VERSION : 0.0
   STRUCT
      doMotorOn : Bool;   // Systemoutput: Status for Motor OFF
      doMotorOff : Bool;   // Systemoutput: Status for Motor ON
      doCycleOn : Bool;   // Systemoutput: Robotprogram is running
      doIRBinAuto : Bool;   // Systemoutput: Robot is in operationmode AUTO
      doSysError : Bool;   // Systemoutput: Robot has an systemerror
      doEmStop_Akt : Bool;   // Systemoutput: Emergencystop at robot is active
      doMot_On_OK : Bool;   // Systemoutput: Automaticstopcicuites are OK
      do01_008 : Bool;   // Spare
      doIRBInHome : Bool;   // Worldzoneoutput: Robot is in Homeposition
      doIRBInMaintP : Bool;   // Worldzoneoutput: Robot is in Maintenanceposition
      doIRBOutRange : Bool;   // Worldzoneoutput: Robot near the end of it´s workingarealimitation
      doIRBOutRangMC : Bool;   // Worldzoneoutput: Robot is out of the mould
      doIRBOutRanMC1 : Bool;   // Worldzoneoutput: Robot is outside the mould carrier 1
      doIRBOutRanMC2 : Bool;   // Worldzoneoutput: Robot is outside the mould carrier 2
      doIRBOutRanMC3 : Bool;   // Worldzoneoutput: Robot is outside the mould carrier 3
      doIRBOutRanMC4 : Bool;   // Worldzoneoutput: Robot is outside the mould carrier 4
      doCycleStarted : Bool;   // The programcycle is startet
      doCycleEnd : Bool;   // The programcycle is finished
      doProgNoReaded : Bool;   // The programnumber is readed
      doShotDigOut : Bool;   // 1st digital Shotware output // Signal to open the mixinghead
      doStopFormPLC : Bool;   // Signal to stop the foaming because the robotprogram has stoped
      doShotBreak : Bool;
      doCloseMould : Bool;   // Signal that the robot is out of the mould
      doCP_forward : Bool;
      doIRBInMaintP2 : Bool;   // Worldzoneoutput: Robot is in 2. Maintenanceposition
      do01_026 : Bool;   // Spare
      doIRBSyncWobj : Bool;   // The robot is synchronized (Tracking)
      doRobWaitWobj : Bool;   // The robot is waiting for synchronizes (Tracking)
      doInPosTeach : Bool;   // The robot is in the position to teaching
      doConveyorStopped : Bool;   // The conveyor is stop
      doZeroSpeed : Bool;   // Systemoutput: Conveyer is not moving
      do01_032 : Bool;   // Spare
      do01_033 : Bool;   // Spare
      doSafetyControlPos : Bool;   // Signal to control the synchronization position
      doSafetySynchronized : Bool;   // Signal from Robot EPS is synchronize
      doSafetySyncSwitch : Bool;   // Signal from Robot sync switch is actuated
      doSafetyArea_1 : Bool;   // 1 Safe Output Safe move / EPS
      doSafetyArea_2 : Bool;   // 2 Safe Output Safe move / EPS
      doSafetyArea_3 : Bool;   // 3 Safe Output Safe move / EPS
      doSafetyArea_4 : Bool;   // 4 Safe Output Safe move / EPS
      doSafetyArea_5 : Bool;   // 5 Safe Output Safe move / EPS
      doSafetyArea_6 : Bool;   // 6 Safe Output Safe move / EPS
      doSafetyArea_7 : Bool;   // 7 Safe Output Safe move / EPS
      doSafetyArea_8 : Bool;   // 8 Safe Output Safe move / EPS
      doSafetyPreWarn : Bool;   // Signal from pre warning robot sync
      doSafeZoneActiv : Bool;   // Robot is inside of a safe tool zone
      do01_047 : Bool;   // Spare
      doClose_Mould_1 : Bool;
      doClose_Mould_2 : Bool;
      doClose_Mould_3 : Bool;
      doClose_Mould_4 : Bool;
      doIRBinSprayP : Bool;
      doSprayValveOn : Bool;
      doStartSpray : Bool;
      doSprayEnd : Bool;
      doInWaitPos : Bool;   // Signal robot is waiting in teh waiting position
      doIRBInWaitP : Bool;   // Signal robot is waiting in teh waiting position // Cube
      do01_058 : Bool;   // Spare
      do01_059 : Bool;   // Spare
      doCleaningPLC : Bool;   // Control the mixinghead cleaner or a brush station
      doCleanOsziJet : Bool;   // Control the air for blow out the oszilation holes
      doBlowAir : Bool;   // Control the air for blow inside the mixinghead
      doCleanBrushOn : Bool;   // Control the cleaning for the mixinghead
      doFlushing : Bool;
      doInFlushposSpray : Bool;
      doShotDigOut2 : Bool;   // 2nd digital Shotware output
      doShotDigOut3 : Bool;   // 3rd digital Shotware output
      do01_068 : Bool;   // Spare
      do01_069 : Bool;   // Spare
      do01_070 : Bool;   // Spare
      do01_071 : Bool;   // Spare
      do01_072 : Bool;   // Spare
      do01_073 : Bool;   // Spare
      do01_074 : Bool;   // Spare
      do01_075 : Bool;   // Spare
      do01_076 : Bool;   // Spare
      do01_077 : Bool;   // Spare
      do01_078 : Bool;   // Spare
      do01_079 : Bool;   // Spare
      do01_080 : Bool;   // Spare
      do10_81_88 : Byte;   // Spare
      goMouldActBit0 : Bool;   // Nummer der Form (1..7) welche zur Zeit bearbeitet wird (Gruppenausgang 0)
      goMouldActBit1 : Bool;   // Nummer der Form (1..7) welche zur Zeit bearbeitet wird (Gruppenausgang 1)
      goMouldActBit2 : Bool;   // Nummer der Form (1..7) welche zur Zeit bearbeitet wird (Gruppenausgang 2)
      go10_92 : Bool;   // Reserve
      go10_93 : Bool;   // Reserve
      go10_94 : Bool;   // Reserve
      go10_95 : Bool;   // Reserve
      go10_96 : Bool;   // Reserve
      GOError : Byte;   // Fehlernummer bei der Bearbeitung des Programms (Gruppenausgang)
      goxFIProgBit0 : Bool;   // Nummer des Faserprogrammes an den Rechner (Gruppenausgang der Shotware, Bit 0)
      goxFIProgBit1 : Bool;   // Nummer des Faserprogrammes an den Rechner (Gruppenausgang der Shotware, Bit 1)
      goxFIProgBit2 : Bool;   // Nummer des Faserprogrammes an den Rechner (Gruppenausgang der Shotware, Bit 2)
      goxFIProgBit3 : Bool;   // Nummer des Faserprogrammes an den Rechner (Gruppenausgang der Shotware, Bit 3)
      go10_117 : Bool;   // Reserve
      go10_118 : Bool;   // Reserve
      go10_119 : Bool;   // Reserve
      go10_120 : Bool;   // Reserve
      goOscixFIBit0 : Bool;   // Bit des Oszillierprogrammes // X1 (2'ter Gruppenausgang der Shotware, Bit 0)
      goOscixFIBit1 : Bool;   // Bit des Oszillierprogrammes // X2 (2'ter Gruppenausgang der Shotware, Bit 1)
      goOscixFIBit2 : Bool;   // Bit des Oszillierprogrammes // Y1 (2'ter Gruppenausgang der Shotware, Bit 2)
      goOscixFIBit3 : Bool;   // Bit des Oszillierprogrammes // Y2 (2'ter Gruppenausgang der Shotware, Bit 3)
      go10_125 : Bool;   // Reserve
      go10_126 : Bool;   // Reserve
      go10_127 : Bool;   // Reserve
      go10_128 : Bool;   // Reserve
   END_STRUCT;
END_TYPE

TYPE "ABB_IRC6_Messages"
VERSION : 0.0
   STRUCT
      Rob_ST_01_16 : Struct
         FLT_No_009 : Bool;
         FLT_No_010 : Bool;
         FLT_No_011 : Bool;
         FLT_No_012 : Bool;
         FLT_No_013 : Bool;
         FLT_No_014 : Bool;
         FLT_No_015 : Bool;
         FLT_No_016 : Bool;
         FLT_No_001 : Bool;
         FLT_No_002 : Bool;
         FLT_No_003 : Bool;
         FLT_No_004 : Bool;
         FLT_No_005 : Bool;
         FLT_No_006 : Bool;
         FLT_No_007 : Bool;
         FLT_No_008 : Bool;
      END_STRUCT;
      Rob_ST_17_32 : Struct
         FLT_No_025 : Bool;   // IRB auf dem Weg zur Form!
         FLT_No_026 : Bool;   // IRB wartet in der Vorposition der Form auf das Sartsignal der SPS!
         FLT_No_027 : Bool;   // IRB in Formträger <X> Formnummer <Y> Teilschuss <Z>
         FLT_No_028 : Bool;   // IRB außerhalb der Form nach dem Schäumen!
         FLT_No_029 : Bool;   // IRB auf dem Weg zum Reinigungsstation!
         FLT_No_030 : Bool;   // IRB ist in der Reinigungsstation! IRB wartet auf das Signal Reinigen starten
         FLT_No_031 : Bool;   // IRB ist in der Reinigungsstation! IRB wartet auf das Signal Reinigen beendet
         FLT_No_032 : Bool;   // IRB auf dem Weg zur Homeposition!
         FLT_No_017 : Bool;
         FLT_No_018 : Bool;
         FLT_No_019 : Bool;   // Falsche Programmnummer!
         FLT_No_020 : Bool;   // Es wurde seit 1h kein Startsignal an den Roboter übermittelt!
         FLT_No_021 : Bool;   // Das Signal <diReadProgNr> von der SPS zum IRB wird nicht zurückgesetzt!
         FLT_No_022 : Bool;   // Der von der SPS übertragene Mouldcode liegt außerhalb des zulässigen Bereiches
         FLT_No_023 : Bool;   // Der von der SPS übertragene Timecode liegt außerhalb des zulässigen Bereiches
         FLT_No_024 : Bool;   // Die aktuelle Schußzeit ist kleiner 1 sec!
      END_STRUCT;
      Rob_ST_33_48 : Struct
         FLT_No_041 : Bool;   // Bitte geben Sie die Formträger- nummer ein auf welcher die Form geteacht wird!
         FLT_No_042 : Bool;   // Starten Sie das Programm nun nur noch Schrittweise!
         FLT_No_043 : Bool;   // Zykluszeit 1 // Zykluszeit 2 // Zykluszeit 3 // Zykluszeit 4
         FLT_No_044 : Bool;   // Fehlerhafte Auswahl des FT! Es wurde kein Werkobjekt zugeordnet!
         FLT_No_045 : Bool;   // Programm wurde gestopt!
         FLT_No_046 : Bool;   // Soll das nächste Werkzeug optimiert werden?
         FLT_No_047 : Bool;   // Der Roboter wartet auf die Syncronisation!
         FLT_No_048 : Bool;   // Sprachauswahl!
         FLT_No_033 : Bool;   // IRB ist in der Homeposition!
         FLT_No_034 : Bool;   // IRB auf dem Weg zur Wartungsposition!
         FLT_No_035 : Bool;   // IRB ist in der Wartungsposition!
         FLT_No_036 : Bool;   // IRB wartet auf <Zyklus-Start> Signal!
         FLT_No_037 : Bool;   // IRB liest Daten von der SPS!
         FLT_No_038 : Bool;   // IRB wartet auf <Schäumen-Start> Signal von der SPS!
         FLT_No_039 : Bool;   // IRB wartet auf <Schäumen-Beenden> Signal von der SPS!
         FLT_No_040 : Bool;   // Bitte geben Sie das zu teachende Programm ein!
      END_STRUCT;
      Rob_ST_49_64 : Struct
         FLT_No_057 : Bool;   // Angewähle Optionen: Shotware: Ja // Tracking : No // Programm Verschiebung: No
         FLT_No_058 : Bool;   // Angewähle Optionen: Shotware: No // Tracking : Ja // Programm Verschiebung: Ja
         FLT_No_059 : Bool;   // Angewähle Optionen: Shotware: No // Tracking : Ja // Programm Verschiebung: No
         FLT_No_060 : Bool;   // Angewähle Optionen: Shotware: No // Tracking : No // Programm Verschiebung: Ja
         FLT_No_061 : Bool;   // Angewähle Optionen: Shotware: No // Tracking : No // Programm Verschiebung: No
         FLT_No_062 : Bool;   // Zum Ändern der Daten benötigen Sie ein Password! Möchten Sie diese Daten ändern
         FLT_No_063 : Bool;   // Bitte geben Sie das Password ein. Password:
         FLT_No_064 : Bool;   // Sie sind nicht berechtigt diese Daten zu ändern!
         FLT_No_049 : Bool;   // Sprachauswahl!
         FLT_No_050 : Bool;   // Sollen die Texte auf dem Bildschirm angezeigt werden?
         FLT_No_051 : Bool;   // Wurde der Roboter mit der Option <SHOTWARE> gebooted?
         FLT_No_052 : Bool;   // Wurde der Roboter mit der Option <Conveyer - Tracking> gebooted?
         FLT_No_053 : Bool;   // Soll das Bewegugsprogram auf einem Formträger verschoben werden?
         FLT_No_054 : Bool;   // Angewähle Optionen: Shotware: Ja // Tracking : Ja // Programm Verschiebung: Ja
         FLT_No_055 : Bool;   // Angewähle Optionen: Shotware: Ja // Tracking : Ja // Programm Verschiebung: No
         FLT_No_056 : Bool;   // Angewähle Optionen: Shotware: Ja // Tracking : No // Programm Verschiebung: Ja
      END_STRUCT;
      Rob_ST_65_80 : Struct
         FLT_No_073 : Bool;
         FLT_No_074 : Bool;
         FLT_No_075 : Bool;
         FLT_No_076 : Bool;
         FLT_No_077 : Bool;
         FLT_No_078 : Bool;
         FLT_No_079 : Bool;
         FLT_No_080 : Bool;
         FLT_No_065 : Bool;   // Geschwindigkeits - Override <100% !!! Soll dieser nun auf 100% gesetzt werden?
         FLT_No_066 : Bool;   // KM-SOFTWARE!!! SIE sind nicht Autorisiert diese Software zu benutzen!
         FLT_No_067 : Bool;   // Bewegungszeit 1 // Bewegungszeit 2 // Bewegungszeit 3 // Bewegungszeit 4
         FLT_No_068 : Bool;   // Starten Sie nun das zu teachende Programm über das Menü Spezial - 4!
         FLT_No_069 : Bool;   // Abbruch Datenlesen von der SPS!
         FLT_No_070 : Bool;
         FLT_No_071 : Bool;
         FLT_No_072 : Bool;
      END_STRUCT;
   END_STRUCT;
END_TYPE

TYPE "IDM_210_Digout_PWM"
VERSION : 0.1
   STRUCT
      Address : Word;
      Active : Bool;
      ChckConnFault : Bool;
      ChckConnDone : Bool;
      Resourcen : Struct
         Request : Bool;
         Transmitting : Bool;
         Active : Bool;
         Data : Struct
            Kanal : Byte;
         END_STRUCT;
      END_STRUCT;
      GeneralParameters : Struct
         Request : Bool;
         Transmitting : Bool;
         Active : Bool;
         Data : Struct
            Periodendauer : DWord;
         END_STRUCT;
      END_STRUCT;
   END_STRUCT;
END_TYPE

TYPE "UDT041_SWU_State"
TITLE = State of switch over units
VERSION : 0.0
   STRUCT
      SWU_OK : Bool;   // Minimum one switch over unit is activated
      Min_1_SWU_release : Bool;   // Minimum one switch over unit is released
      Open_SWU_disabelt : Bool;   // The actual SWU using for recirculation was disabelt
      Hubcounter_OK : Bool;   // The amount of shot hubs was reached
      Switchingtime_runs : Bool;   // Time after switch over SWU running
      Stoptime_runs : Bool;   // Time after switch off SWU running
      SWU_not_released : Bool;   // The requested SWU not released
      Spare_0_7 : Bool;
      FLT_open_SWU_disabelt : Bool;   // Fault selected switch over unit disabelt
      FLT_No_SWU_selected : Bool;   // Fault no switch over unit selected
      FLT_Sel_SWU_not_released : Bool;   // Fault selected switch over unit not released
      FaultLevel_1 : Bool;   // A fault group 1 exists
      FaultLevel_2 : Bool;   // A fault group 2 exists
      FaultLevel_3 : Bool;   // A fault group 3 exists
      CycleStarted : Bool;   // A cycle was started and is still running
      Spare_1_7 : Bool;
      ActualSWU : Int;   // No of actual open SWU
      SWU_for_Circulation : DWord;   // Buffer of actual SWU during recirculation
      SWU_released : "UDT001_DWord_1_32";   // Bitarea of released SWU
      Target_SWU : "UDT001_DWord_1_32";   // Bitarea witch released SWU will be actvated
      Open_SWU : "UDT001_DWord_1_32";   // Bitarea witch released SWU is activated
      Open_SWU_allone : "UDT001_DWord_1_32";   // Bitarea of the "alone" activated SWU
   END_STRUCT;
END_TYPE

TYPE "UDT042_MH_Select"
TITLE = State of activated and selected mixingheads
VERSION : 0.0
   STRUCT
      Release_MH : "UDT001_DWord_1_32";
      Mixingheadvalve : "UDT001_DWord_1_32";
      Shotcounter : "UDT001_DWord_1_32";
      Countervalue : Word;
      Counterrampe : Bool;
      ImpCounterOn : Bool;   // Impuls to count one value additional
      Spare_14_2 : Bool;
      Spare_14_3 : Bool;
      Spare_14_4 : Bool;
      Spare_14_5 : Bool;
      Spare_14_6 : Bool;
      Spare_14_7 : Bool;
      Cleaningpiston_OK : Bool;
      Spare_15_1 : Bool;
      Spare_15_2 : Bool;
      Spare_15_3 : Bool;
      Spare_15_4 : Bool;
      Spare_15_5 : Bool;
      Spare_15_6 : Bool;
      Spare_15_7 : Bool;
   END_STRUCT;
END_TYPE

TYPE "IDM_212_Digout_Oscillation"
VERSION : 0.1
   STRUCT
      Address : Int;
      Active : Bool;
      ChckConnFault : Bool;
      ChckConnDone : Bool;
      Resourcen : Struct
         Request : Bool;
         Transmitting : Bool;
         Active : Bool;
         Data : Struct
            Kanal : Struct
               Bit0 : Bool;
               Bit1 : Bool;
               Bit2 : Bool;
               Bit3 : Bool;
               Bit4 : Bool;
               Bit5 : Bool;
               Bit6 : Bool;
               Bit7 : Bool;
            END_STRUCT;
         END_STRUCT;
      END_STRUCT;
      GeneralParameters : Struct
         Request : Bool;
         Transmitting : Bool;
         Active : Bool;
         Data : Struct
            Einschaltdauer : Bool;
            "Symmetrie X" : Bool;
            "Symmetrie Y" : Bool;
            Phasenverschiebung : Bool;
         END_STRUCT;
      END_STRUCT;
   END_STRUCT;
END_TYPE

TYPE "IDM_301_Analogin_Default"
VERSION : 0.1
   STRUCT
      Address : Word;
      Active : Bool;
      ChckConnFault : Bool;
      ChckConnDone : Bool;
      Skalierung : Struct
         Request : Bool;
         Transmitting : Bool;
         Active : Bool;
         Data : Struct
            Bereichsobergrenze : Int := 10000;
            Bereichsuntergrenze : Int := -10000;
         END_STRUCT;
      END_STRUCT;
      Filterung : Struct
         Request : Bool;
         Transmitting : Bool;
         Active : Bool;
         Data : Struct
            Mittelwertzeit : Int := 100;
         END_STRUCT;
      END_STRUCT;
      Grenzen : Struct
         Request : Bool;
         Transmitting : Bool;
         Active : Bool;
         Data : Struct
            ObererGrenzwert : Int := 5000;
            UntererGrenzwert : Int;
            AuslösezeitObererGrenzwert : Int := 100;
            ErholungszeitObererGrenzwert : Int := 100;
            AuslösezeitUntererGrenzwert : Int := 100;
            ErholungszeitUntererGrenzwert : Int := 100;
         END_STRUCT;
      END_STRUCT;
   END_STRUCT;
END_TYPE

TYPE "UDT045_Nozzlecontrol"
TITLE = State MH-Nozzle
VERSION : 0.1
   STRUCT
      Select_RCL_to_Nozzle : Bool;
      Select_RCL_not_to_Nozzle : Bool;
      Spare_02 : Bool;
      Spare_03 : Bool;
      Spare_04 : Bool;
      Spare_05 : Bool;
      Spare_06 : Bool;
      Spare_07 : Bool;
      Spare_10 : Bool;
      Spare_11 : Bool;
      Spare_12 : Bool;
      Spare_13 : Bool;
      Spare_14 : Bool;
      Spare_15 : Bool;
      Spare_16 : Bool;
      Spare_17 : Bool;
   END_STRUCT;
END_TYPE

TYPE "UDT046_MH_Lock"
TITLE = State locking of a mixinghead at a mould carrier
VERSION : 0.1
   STRUCT
      Switch_MH_Lock_ON_OFF : Bool;
      MH_Locked : Bool;   // Mixinghead locked do not move
      MH_UnLocked : Bool;   // Mixinghead unlocked mixinghead can be moved
      ReleaseUnlockAfterShot : Bool;
      MH_Lock_active : Bool;
      HF_MH_Unlocked : Bool;
      FL_MH_Unlocked : Bool;   // Flag mixinghead unlocked
      ShotRelease : Bool;   // Shot release after locking
      Fault_RT_Lock : Bool;   // Time locking mixinghead takes too long
      Fault_RT_Unlock : Bool;   // Time unlocking mixinghead takes too long
      FaultLevel_1 : Bool;   // A fault group 1 exist
      FaultLevel_2 : Bool;   // A fault group 2 exist
      FaultLevel_3 : Bool;   // A fault group 3 exist
      Spare15 : Bool;
      Spare16 : Bool;
      Spare17 : Bool;
      Spare : Int;
      State_MHLock : Int;   // 1: locked; 2: faulty; 3:locking required but still unlocked
   END_STRUCT;
END_TYPE

TYPE "IDM_302_Analogin_Default_8"
VERSION : 0.1
   STRUCT
      Address : Int;
      Active : Bool;
      ChckConnFault : Bool;
      ChckConnDone : Bool;
      X14_0 : Struct
         Request : Bool;
         Transmitting : Bool;
         Active : Bool;
         Data : Struct
            "Data[1]" : Struct
               Betriebsart : Byte;
               Reserve : Byte;
               Bereichsobergrenze : Int := 1000;
               Bereichsuntergrenze : Int := 0;
               Mittelwertzeit : Int := 100;
            END_STRUCT;
            "Data[2]" : Struct
               Betriebsart : Byte;
               Reserve : Byte;
               Bereichsobergrenze : Int := 1000;
               Bereichsuntergrenze : Int := 0;
               Mittelwertzeit : Int := 100;
            END_STRUCT;
            "Data[3]" : Struct
               Betriebsart : Byte;
               Reserve : Byte;
               Bereichsobergrenze : Int := 1000;
               Bereichsuntergrenze : Int := 0;
               Mittelwertzeit : Int := 100;
            END_STRUCT;
            "Data[4]" : Struct
               Betriebsart : Byte;
               Reserve : Byte;
               Bereichsobergrenze : Int := 1000;
               Bereichsuntergrenze : Int := 0;
               Mittelwertzeit : Int := 100;
            END_STRUCT;
            "Data[5]" : Struct
               Betriebsart : Byte;
               Reserve : Byte;
               Bereichsobergrenze : Int := 1000;
               Bereichsuntergrenze : Int := 0;
               Mittelwertzeit : Int := 100;
            END_STRUCT;
            "Data[6]" : Struct
               Betriebsart : Byte;
               Reserve : Byte;
               Bereichsobergrenze : Int := 1000;
               Bereichsuntergrenze : Int := 0;
               Mittelwertzeit : Int := 100;
            END_STRUCT;
            "Data[7]" : Struct
               Betriebsart : Byte;
               Reserve : Byte;
               Bereichsobergrenze : Int := 1000;
               Bereichsuntergrenze : Int := 0;
               Mittelwertzeit : Int := 100;
            END_STRUCT;
            "Data[8]" : Struct
               Betriebsart : Byte;
               Reserve : Byte;
               Bereichsobergrenze : Int := 1000;
               Bereichsuntergrenze : Int := 0;
               Mittelwertzeit : Int := 100;
            END_STRUCT;
         END_STRUCT;
      END_STRUCT;
   END_STRUCT;
END_TYPE

TYPE "IDM_401_Analogout_Default"
VERSION : 0.1
   STRUCT
      Address : Int;
      Active : Bool;
      ChckConnFault : Bool;
      ChckConnDone : Bool;
      GeneralParameters : Struct
         Request : Bool;
         Transmitting : Bool;
         Active : Bool;
         Data : Struct
            Ausgangskanal : Struct
               Bit0 : Bool;
               Bit1 : Bool;
               Bit2 : Bool;
               Spare3 : Bool;
               Spare4 : Bool;
               Spare5 : Bool;
               Spare6 : Bool;
               Spare7 : Bool;
               Bereichsobergrenze : Int := 10000;   // 1000..32767
               Bereichsuntergrenze : Int := -10000;   // -32767..32767
               Rampenzeit : Int := 1000;   // 1..5000
            END_STRUCT;
         END_STRUCT;
      END_STRUCT;
   END_STRUCT;
END_TYPE

TYPE "IDM_402_Analogout_Flow_Controller"
VERSION : 0.1
   STRUCT
      Address : Word;
      Active : Bool;
      ChckConnFault : Bool;
      ChckConnDone : Bool;
      GeneralParameters : Struct
         Request : Bool;
         Transmitting : Bool;
         Active : Bool;
         Data : Struct
            Kalibrierfaktor : DInt := 10000;   // 100..4294967295*0.0001g/Puls
            MaxDurchfluss : DInt := 1000;   // 100..4294967295*0.01g/s
            Nachstellzeit : Int := 50;   // 1..10000ms
            Filterzeit : Int := 200;   // 1..1024
         END_STRUCT;
      END_STRUCT;
      Grenzen : Struct
         Request : Bool;
         Transmitting : Bool;
         Active : Bool;
         Data : Struct
            ObergrenzeStellgröße : Int := 10000;   // 0..10000
            UntergrenzeStellgröße : Int := 0;   // -10000..10000
            VerzögerungAlarmObergrenze : Int := 1000;   // 1..10000ms
            VerzögerungAlarmUntergrenze : Int := 1000;   // 1..10000ms
         END_STRUCT;
      END_STRUCT;
      SkalierungAI : Struct
         Request : Bool;
         Transmitting : Bool;
         Active : Bool;
         Data : Struct
            Bereichsobergrenze : Int := 10000;   // 0..32767
            Bereichsuntergrenze : Int := -10000;   // -32767..32767
            Mittelwertzeit : Int := 100;   // 1..1000ms
         END_STRUCT;
      END_STRUCT;
   END_STRUCT;
END_TYPE

TYPE "IDM_415_Analogout_Flow_Controller_Float"
VERSION : 0.1
   STRUCT
      Address : Int;
      Active : Bool;
      ChckConnFault : Bool;
      ChckConnDone : Bool;
      "I/O" : Struct
         InputData : Struct
            Flow : Real;
            Weight : Real;
            ActPresSDA : Int;
            Control : Struct
               ZeroFlow : Bool;   // Durchfluss ist Null
               SDAactiv : Bool;   // SDA ist aktiv
               FlowControlUpperLimit : Bool;   // Durchflussregler arbeit an der Obergrenze
               FlowControlLowerLimit : Bool;   // Durchflussregler arbeit an der Untergrenze
               FlowLowerLimit : Bool;   // Tatsächlicher Durchfluss ist unter der Toleranzgrenze
               FlowUpperLimit : Bool;   // Tatsächlicher Durchfluss ist über der Toleranzgrenze
               Spare06 : Bool;
               Spare07 : Bool;
            END_STRUCT;
         END_STRUCT;
         OutputData : Struct
            Flow : Real;
            FlowSDA : Real;
            PressSDA : Real;
            actPressSDA : Real;
            Control : Struct
               NonControledValue : Bool;   // Gesteuerte Werte ausgeben
               ControledValue : Bool;   // Geregelte Werte ausgeben
               SetValueOverlay : Bool;   // Sollwertüberlagerung
               SDATrig : Bool;   // SDA triggern
               ResetWeight : Bool;   // Gewicht zurücksetzen
               Spare05 : Bool;
               Spare06 : Bool;
               Spare07 : Bool;
            END_STRUCT;
         END_STRUCT;
      END_STRUCT;
      Hardware : Struct
         Request : Bool;
         Transmitting : Bool;
         Active : Bool;
         Data : Struct
            AO_Ausgangskanal_FU : Byte;
            AI_Eingangskanal_Druck : Byte;
            DI_Eingangskanal_Puls : Byte;
            Konfig1 : Byte;
            Konfig2 : Byte;
            Rampenzeit : Real := 0.1;   // 0.001..5.000
         END_STRUCT;
      END_STRUCT;
      GeneralParameters : Struct
         Request : Bool;
         Transmitting : Bool;
         Active : Bool;
         Busy : Bool;
         Done : Bool;
         Data : Struct
            Kalibrierfaktor : Real := 1.0;   // 0.01..429496.72 g/Puls
            MaxDurchfluss : Real := 100.0;   // 1..42949672.0 g/s
            Nachstellzeit : Real := 0.05;   // 0.001..10s
            Filterzeit : Real := 0.2;   // 0.001..1.024s
         END_STRUCT;
      END_STRUCT;
      Grenzen : Struct
         Request : Bool;
         Tranmitting : Bool;
         Active : Bool;
         Busy : Bool;
         Done : Bool;
         Data : Struct
            ObergrenzeStellgröße : Real := 1.0;   // 0..1s
            UntergrenzeStellgröße : Real := 0.0;   // -1..1s
            VerzögerungAlarmObergrenze : Real := 1.0;   // 0.001..10s
            VerzögerungAlarmUntergrenze : Real := 1.0;   // 0.001..10s
         END_STRUCT;
      END_STRUCT;
      SkalierungAI : Struct
         Request : Bool;
         Transmitting : Bool;
         Active : Bool;
         Busy : Bool;
         Done : Bool;
         Data : Struct
            Bereichsobergrenze : Real := 600.0;   // 100..32767
            Bereichsuntergrenze : Real := 0.0;   // -32767..32767
            Mittelwertzeit : Real := 0.1;   // 0.001..1s
         END_STRUCT;
      END_STRUCT;
      Visualisierung : Struct
         BetriebsartAnalogausgang : Byte;   // Byte 0 Bit 0-2
         BipolarerAusgang : Byte;   // Byte 0 Bit 3
         Polarität : Byte;   // Byte 0 Bit 4
         BetriebsartAnalogeingang : Byte;   // Byte 0 Bit 5-7
         BetriebsartQuadraturdekoder : Byte;   // Byte 1 Bit 0-1
         QuelleIstdruck : Byte;   // Byte 1 Bit 2
         Dichte : Real;
      END_STRUCT;
   END_STRUCT;
END_TYPE

TYPE "IDM_501_Analogin_Temperature"
VERSION : 0.1
   STRUCT
      Address : Word;
      Active : Bool;
      ChckConnFault : Bool;
      ChckConnDone : Bool;
      X12_0 : Struct
         Request : Bool;
         Transmitting : Bool;
         Active : Bool;
         Data : Struct
            Mittelwertzeit : Int := 100;
            ErsatzwertDrahtbruch : Bool;
            Bits : Struct
               B0_Einheit : Bool;
               B1_Einheit : Bool;
               B2 : Bool;
               B3 : Bool;
               B4 : Bool;
               B5 : Bool;
               B6 : Bool;
               B7 : Bool;
            END_STRUCT;
         END_STRUCT;
      END_STRUCT;
   END_STRUCT;
END_TYPE

TYPE "IDM_502_Analogin_Temperature_8"
VERSION : 0.1
   STRUCT
      Address : Int;
      Active : Bool;
      ChckConnFault : Bool;
      ChckConnDone : Bool;
      TemperatureInput : Struct
         Request : Bool;
         Transmitting : Bool;
         Active : Bool;
         Data : Array[1..8] of Struct
            Mittelwertzeit : Int;
            ErsatzwertDrahtbruch : Int;
            Einheit : Byte;
            Reserve : Byte;
         END_STRUCT;
      END_STRUCT;
   END_STRUCT;
   // TemperatureInput.Data[1].Mittelwertzeit := 100;
   // TemperatureInput.Data[2].Mittelwertzeit := 100;
   // TemperatureInput.Data[3].Mittelwertzeit := 100;
   // TemperatureInput.Data[4].Mittelwertzeit := 100;
   // TemperatureInput.Data[5].Mittelwertzeit := 100;
   // TemperatureInput.Data[6].Mittelwertzeit := 100;
   // TemperatureInput.Data[7].Mittelwertzeit := 100;
   // TemperatureInput.Data[8].Mittelwertzeit := 100;
END_TYPE

TYPE "UDT053_Pump"
TITLE = State of a metering pump
VERSION : 0.0
   STRUCT
      FLT_Exist : Bool;   // A fault exist
      FaultLevel_1 : Bool;   // A fault group 1 exist
      FaultLevel_2 : Bool;   // A fault group 2 exist
      FaultLevel_3 : Bool;   // A fault group 3 exist
      High_rpm : Bool;   // Request to drive component pump in high speed
      Metering_to_PUC : Bool;   // Request of metering the component
      Selection_Feedingpump : Bool;   // Request to start the feed pump
      Main_Pumpselection : Bool;   // Request to start the component pump
      Netrelais : Bool;   // Request to switch the main conactor of the component pump
      Controllrelease_to_FC : Bool;   // Activation of the control release of the frequence unit of the component
      Enableclosedloop : Bool;   // PLC-release to control the component flow at modul
      Valve_2_point_selection : Bool;   // Activate the valve of the 2-point adjustment of component
      Release_Startup_FC : Bool;   // Delay to switch ON frequence unit after power lost or emergency stop
      Puls_SDA : Bool;   // Flag of the signal to switch over to the quick pressure build up
      Rampe_Voltage_Off : Bool;   // Flag of delay to switch ON after power lost
      Start_Startupdelay : Bool;   // Information that delay time to switch ON after power lost is running
      IntervalPause : Bool;   // Pause time if interval mode is running
      Ventingtime_finished : Bool;   // The ventilation time is over
      Net_Ventilation : Bool;   // Activation of ventilation pump
      FLT_Ventilation : Bool;   // Fault: Motorprotection ventilation drive of drive pump
      Mes_PumpDeselected : Bool;   // Message: Pump is deselected for maintenance purposes
      Mes_PumpDeselectedInt : Bool;   // Message: Pump is deselected and runs in interval mode
      FLT_MotorFan : Bool;   // Fault: Motorprotection external fan of motor
      HF_FPPumpDeselectedInt : Bool;   // Flag Pump is deselected and runs in interval mode
      "2PointAdjustmentSelected" : Bool;
      Block_is_active : Bool;   // The program block passed through // Info at least one component is active
   END_STRUCT;
END_TYPE

TYPE "IDM_601_Mixinghead_Digital"
VERSION : 0.1
   STRUCT
      Address : Int;
      Active : Bool;
      ChckConnFault : Bool;
      ChckConnDone : Bool;
      GeneralParameters : Struct
         Request : Bool;
         Transmitting : Bool;
         Active : Bool;
         Data : Struct
            EingangskanalMK_Ini : Byte;   // 0..32
            EingangskanalFreigabe : Byte;   // 0..32
            Ventilausgang : Byte;   // 0..31
            MischkopfKanal : Byte;   // 0..3
         END_STRUCT;
      END_STRUCT;
      Zeiten : Struct
         Request : Bool;
         Transmitting : Bool;
         Active : Bool;
         Data : Struct
            ÜberwachungszeitÖffnen : Real;   // 1..32000ms
            ÜberwachungszeitSchließen : Real;   // 1..32000ms
            ErlaubtePrellzeit : Real;   // 0..100
         END_STRUCT;
      END_STRUCT;
      Zeiten_2 : Struct
         Request : Bool;
         Transmitting : Bool;
         Active : Bool;
         Data : Struct
            Verzögerungszeit_HW_Freigabe : Real;   // 1..32000ms
         END_STRUCT;
      END_STRUCT;
   END_STRUCT;
END_TYPE

TYPE "IDM_605_Mixinghead_Analog"
VERSION : 0.1
   STRUCT
      Address : Int;
      Active : Bool;
      ChckConnFault : Bool;
      ChckConnDone : Bool;
      Resourcen : Struct
         Request : Bool;
         Transmitting : Bool;
         Active : Bool;
         Data : Struct
            EingangskanalMK_Ini : Struct
               Bool0 : Bool;
               Bool1 : Bool;
               Bool2 : Bool;
               Bool3 : Bool;
               Bool4 : Bool;
               Bool5 : Bool;
               Spare6 : Bool;
               Spare7 : Bool;
            END_STRUCT;
            EingangskanalFreigabe : Struct
               Bool0 : Bool;
               Bool1 : Bool;
               Bool2 : Bool;
               Bool3 : Bool;
               Bool4 : Bool;
               Bool5 : Bool;
               Bool6 : Bool;
               Bool7 : Bool;
            END_STRUCT;
            AnalogerAusgang : Struct
               Bool0 : Bool;
               Bool1 : Bool;
               Bool2 : Bool;
               Spare3 : Bool;
               Spare4 : Bool;
               Spare5 : Bool;
               Spare6 : Bool;
               Spare7 : Bool;
            END_STRUCT;
            Betriebsart : Struct
               Bool0 : Bool;
               Bool1 : Bool;
               Bool2 : Bool;
               Spare3 : Bool;
               Spare4 : Bool;
               Spare5 : Bool;
               Spare6 : Bool;
               Spare7 : Bool;
            END_STRUCT;
            MischkopfKanal : Struct
               Bool0 : Bool;
               Bool1 : Bool;
               Spare2 : Bool;
               Spare3 : Bool;
               Spare4 : Bool;
               Spare5 : Bool;
               Spare6 : Bool;
               Spare7 : Bool;
            END_STRUCT;
         END_STRUCT;
      END_STRUCT;
      Zeiten : Struct
         Request : Bool;
         Transmitting : Bool;
         Active : Bool;
         Data : Struct
            ÜberwachungszeitÖffnen : Int := 500;   // 1..32000ms
            ÜberwachungszeitSchließen : Int := 500;   // 1..32000ms
            ErlaubtePrellzeit : Int := 20;   // 0..100
         END_STRUCT;
      END_STRUCT;
      Skalierung : Struct
         Request : Bool;
         Transmitting : Bool;
         Active : Bool;
         Data : Struct
            Bereichsobergrenze : Int := 10000;   // 1000..32767
            Bereichsuntergrenze : Int := -10000;   // -32767..32767
         END_STRUCT;
      END_STRUCT;
      StufenAktivierung : Struct
         Request : Bool;
         Transmitting : Bool;
         Active : Bool;
         Data : Struct
            DauerStufe1 : Int := 10;   // 1..32000ms
            DauerStufe2 : Int := 10;   // 1..32000ms
            DauerStufe3 : Int := 10;   // 1..32000ms
            DauerStufe4 : Int := 10;   // 1..32000ms
            DauerStufe5 : Int := 10;   // 1..32000ms
            LevelStufe1 : Int := 10000;   // -32768..1000
            LevelStufe2 : Int := 5000;   // -32768..1000
            LevelStufe3 : Int := 1500;   // -32768..1000
            LevelStufe4 : Int := 500;   // -32768..1000
            LevelStufe5 : Int := 0;   // -32768..1000
         END_STRUCT;
      END_STRUCT;
      StufenRückkehr : Struct
         Request : Bool;
         Transmitting : Bool;
         Active : Bool;
         Data : Struct
            DauerStufe1 : Int := 10;   // 1..32000ms
            DauerStufe2 : Int := 10;   // 1..32000ms
            DauerStufe3 : Int := 10;   // 1..32000ms
            DauerStufe4 : Int := 10;   // 1..32000ms
            DauerStufe5 : Int := 10;   // 1..32000ms
            LevelStufe1 : Int := -10000;   // -32768..1000
            LevelStufe2 : Int := -5000;   // -32768..1000
            LevelStufe3 : Int := -1500;   // -32768..1000
            LevelStufe4 : Int := -500;   // -32768..1000
            LevelStufe5 : Int := 0;   // -32768..1000
         END_STRUCT;
      END_STRUCT;
   END_STRUCT;
END_TYPE

TYPE "IDM_610_CleaningPiston_Digital"
VERSION : 0.1
   STRUCT
      Address : Int;
      Active : Bool;
      ChckConnFault : Bool;
      ChckConnDone : Bool;
      GeneralParameters : Struct
         Request : Bool;
         Transmitting : Bool;
         Active : Bool;
         Data : Struct
            EingangskanalRK_Ini : Byte;   // 0..32
            AusgangRKVentil : Byte;   // 0..31
            MischkopfKanal : Byte;   // 0..3
         END_STRUCT;
      END_STRUCT;
      Zeiten : Struct
         Request : Bool;
         Transmitting : Bool;
         Active : Bool;
         Data : Struct
            ÜberwachungszeitVorfahren : Real := 0.5;   // 1..32000ms
            ÜberwachungszeitRückfahren : Real := 0.5;   // 1..32000ms
            ErlaubtePrellzeit : Real := 0.02;   // 0..100
            WartezeitVorne : Real := 0.5;   // 0..40000000000
            VerzögerungNachSchuss : Real := 0.5;   // 0..40000000000
         END_STRUCT;
      END_STRUCT;
   END_STRUCT;
END_TYPE

TYPE "IDM_615_CleaningPiston_Analog"
VERSION : 0.1
   STRUCT
      Address : Int;
      Active : Bool;
      ChckConnFault : Bool;
      ChckConnDone : Bool;
      GeneralParameters : Struct
         Request : Bool;
         Transmitting : Bool;
         Active : Bool;
         Data : Struct
            EingangskanalRK_Ini : Struct
               Bool0 : Bool;
               Bool1 : Bool;
               Bool2 : Bool;
               Bool3 : Bool;
               Bool4 : Bool;
               Bool5 : Bool;
               Spare6 : Bool;
               Spare7 : Bool;
            END_STRUCT;
            AnalogerAusgang : Struct
               Bool0 : Bool;
               Bool1 : Bool;
               Bool2 : Bool;
               Spare3 : Bool;
               Spare4 : Bool;
               Spare5 : Bool;
               Spare6 : Bool;
               Spare7 : Bool;
            END_STRUCT;
            Betriebsart : Struct
               Bool0 : Bool;
               Bool1 : Bool;
               Bool2 : Bool;
               Spare3 : Bool;
               Spare4 : Bool;
               Spare5 : Bool;
               Spare6 : Bool;
               Spare7 : Bool;
            END_STRUCT;
            MischkopfKanal : Struct
               Bool0 : Bool;
               Bool1 : Bool;
               Spare2 : Bool;
               Spare3 : Bool;
               Spare4 : Bool;
               Spare5 : Bool;
               Spare6 : Bool;
               Spare7 : Bool;
            END_STRUCT;
            Rampenzeit : Int := 1000;   // 1..5000
         END_STRUCT;
      END_STRUCT;
      Zeiten : Struct
         Request : Bool;
         Transmitting : Bool;
         Active : Bool;
         Data : Struct
            ÜberwachungszeitVorfahren : Int := 500;   // 1..32000ms
            ÜberwachungszeitRückfahren : Int := 500;   // 1..32000ms
            ErlaubtePrellzeit : Int := 20;   // 0..100
            WartezeitVorne : Real := 1.0;   // 0..4000000000000
            WartezeitHinten : Real := 1.0;   // 0..4000000000000
         END_STRUCT;
      END_STRUCT;
      Skalierung : Struct
         Request : Bool;
         Transmitting : Bool;
         Active : Bool;
         Data : Struct
            Bereichsobergrenze : Int := 10000;   // 1000..32767
            Bereichsuntergrenze : Int := -10000;   // -32767..32767
         END_STRUCT;
      END_STRUCT;
      StufenAktivierung : Struct
         Request : Bool;
         Transmitting : Bool;
         Active : Bool;
         Data : Struct
            DauerStufe1 : Int := 10;   // 1..32000ms
            DauerStufe2 : Int := 10;   // 1..32000ms
            DauerStufe3 : Int := 10;   // 1..32000ms
            DauerStufe4 : Int := 10;   // 1..32000ms
            DauerStufe5 : Int := 10;   // 1..32000ms
            LevelStufe1 : Int := 10000;   // 0..32767
            LevelStufe2 : Int := 5000;   // 0..32767
            LevelStufe3 : Int := 1500;   // 0..32767
            LevelStufe4 : Int := 500;   // 0..32767
            LevelStufe5 : Int := 0;   // 0..32767
         END_STRUCT;
      END_STRUCT;
      StufenRückkehr : Struct
         Request : Bool;
         Transmitting : Bool;
         Active : Bool;
         Data : Struct
            DauerStufe1 : Int := 10;   // 1..32000ms
            DauerStufe2 : Int := 10;   // 1..32000ms
            DauerStufe3 : Int := 10;   // 1..32000ms
            DauerStufe4 : Int := 10;   // 1..32000ms
            DauerStufe5 : Int := 10;   // 1..32000ms
            LevelStufe1 : Int := -10000;   // -32768..1000
            LevelStufe2 : Int := -5000;   // -32768..1000
            LevelStufe3 : Int := -1500;   // -32768..1000
            LevelStufe4 : Int := -500;   // -32768..1000
            LevelStufe5 : Int := 0;   // -32768..1000
         END_STRUCT;
      END_STRUCT;
   END_STRUCT;
END_TYPE

TYPE "IDM_616_CleaningPiston_Analog_Loop"
VERSION : 0.1
   STRUCT
      Address : Int;
      Active : Bool;
      ChckConnFault : Bool;
      ChckConnDone : Bool;
      GeneralParameters : Struct
         Request : Bool;
         Transmitting : Bool;
         Active : Bool;
         Data : Struct
            AnalogerAusgang : Struct
               Bool0 : Bool;
               Bool1 : Bool;
               Bool2 : Bool;
               Spare3 : Bool;
               Spare4 : Bool;
               Spare5 : Bool;
               Spare6 : Bool;
               Spare7 : Bool;
            END_STRUCT;
            Betriebsart : Struct
               Bool0 : Bool;
               Bool1 : Bool;
               Bool2 : Bool;
               Spare3 : Bool;
               Spare4 : Bool;
               Spare5 : Bool;
               Spare6 : Bool;
               Spare7 : Bool;
            END_STRUCT;
            AnalogerEingang : Struct
               Bool0 : Bool;
               Bool1 : Bool;
               Bool2 : Bool;
               Spare3 : Bool;
               Spare4 : Bool;
               Spare5 : Bool;
               Spare6 : Bool;
               Spare7 : Bool;
            END_STRUCT;
            Betriebsart_1 : Struct
               Bool0 : Bool;
               Bool1 : Bool;
               Spare2 : Bool;
               Spare3 : Bool;
               Spare4 : Bool;
               Spare5 : Bool;
               Spare6 : Bool;
               Spare7 : Bool;
            END_STRUCT;
            MischkopfKanal : Struct
               Bool0 : Bool;
               Bool1 : Bool;
               Spare2 : Bool;
               Spare3 : Bool;
               Spare4 : Bool;
               Spare5 : Bool;
               Spare6 : Bool;
               Spare7 : Bool;
               AnalogerAusgang : Struct
                  Bool0 : Bool;
                  Bool1 : Bool;
                  Bool2 : Bool;
                  Spare3 : Bool;
                  Spare4 : Bool;
                  Spare5 : Bool;
                  Spare6 : Bool;
                  Spare7 : Bool;
               END_STRUCT;
            END_STRUCT;
         END_STRUCT;
      END_STRUCT;
      Zeiten : Struct
         Request : Bool;
         Transmitting : Bool;
         Active : Bool;
         Data : Struct
            ÜberwachungszeitVorfahren : Int := 500;   // 1..32000ms
            ÜberwachungszeitRückfahren : Int := 500;   // 1..32000ms
            WartezeitVorne : Real := 1.0;   // 0..4000000000000
            WartezeitHinten : Real := 1.0;   // 0..4000000000000
            KolbenrückzugVorSchussende : Int := 500;   // 0..32000
         END_STRUCT;
      END_STRUCT;
      Skalierung : Struct
         Request : Bool;
         Transmitting : Bool;
         Active : Bool;
         Data : Struct
            Bereichsobergrenze : Int := 10000;   // 1000..32767
            Bereichsuntergrenze : Int := -10000;   // -32767..32767
         END_STRUCT;
      END_STRUCT;
      Regelparameter : Struct
         Request : Bool;
         Transmitting : Bool;
         Active : Bool;
         Data : Struct
            P_Faktor : Real := 1.0;
            Integrationszeit : Real := 1000.0;
            Differenzierzeit : Real := 0.001;
         END_STRUCT;
      END_STRUCT;
   END_STRUCT;
END_TYPE

TYPE "IDM_620_Mixinghead_NozzleBypass"
VERSION : 0.1
   STRUCT
      Address : Int;
      Active : Bool;
      ChckConnFault : Bool;
      ChckConnDone : Bool;
      Channel : Struct
         Request : Bool;
         Transmitting : Bool;
         Active : Bool;
         Data : Struct
            Konfig1 : Byte;
            Konfig2 : Byte;
            Konfig3 : Byte;
         END_STRUCT;
      END_STRUCT;
      Zeiten : Struct
         Request : Bool;
         Transmitting : Bool;
         Active : Bool;
         Data : Struct
            ÜberlappungD_B : Real := 0.2;   // -32.000..32.000
            ÜberlappungB_D : Real := 0.2;   // -32.000..32.000
            VerzögerungSchussstart : Real := 1.0;   // -32.000..32.000
            VerzögerungSchussende : Real := 1.0;   // -32.000..32.000
         END_STRUCT;
      END_STRUCT;
      Visualisierung : Struct
         OutputForNozzle : Byte;   // 0..32
         PolarityNozzle : Byte;   // 0..1
         OutputForBypass : Byte;   // 0..32
         PolarityBypass : Byte;   // 0..1
         MHChannel : Byte;   // 0..3
      END_STRUCT;
   END_STRUCT;
END_TYPE

TYPE "SZL-IDW#16#xy96_DataSet"
VERSION : 0.1
   STRUCT
      LogicalAddr : Word;
      System : Word;
      API : DWord;
      Station : Word;
      Slot : Word;
      Subslot : Word;
      Offset : Word;
      SetType : Struct
         Herstellernummer : Word;
         Geraet : Word;
         LaufendeNummer : Word;
         ModulIdentifikation1 : Word;
         ModulIdentifikation2 : Word;
         SubmodulIdentifikation1 : Word;
         Submodulidentifikation2 : Word;
      END_STRUCT;
      SetType_UnEqual_ActualType : Array[0..15] of Bool;
      res : Word;
      IOStat : Struct
         BaugruppeWartungsbedarf : Bool;
         BaugruppeWartungsanforderung : Bool;
         res10 : Bool;
         res11 : Bool;
         res12 : Bool;
         res13 : Bool;
         res14 : Bool;
         res15 : Bool;
         BaugruppeGestoert : Bool;
         BaugruppeVorhanden : Bool;
         BaugruppeNichtVerfuegbar : Bool;
         BaugruppeDeaktiviert : Bool;
         StoerungDerStation : Bool;
         M7_BaugruppeHostFuerSup : Bool;   // Baugruppe kann Host für Submodule sein
         res6 : Bool;
         BaugruppeImLokalbussegment : Bool;
      END_STRUCT;
      AreaID_ModuleWidth : Word;
      res_1 : Word;
      res_2 : Word;
      res_3 : Word;
      res_4 : Word;
      res_5 : Word;
      res_6 : Word;
      res_7 : Word;
      res_8 : Word;
      res_9 : Word;
      res_10 : Word;
   END_STRUCT;
END_TYPE

TYPE "UDT061_Cylinder_Manager"
TITLE = State of cylinder Manager
VERSION : 0.0
   STRUCT
      Stop_to_Pause : Bool;   // Request to stop piston in pause position
      All_cylinder_up : Bool;   // All pistons of the plant are at upper end postion
      Spare_0_2 : Bool;
      Spare_0_3 : Bool;
      Spare_0_4 : Bool;
      FlagPistonUp : Bool;   // Edgeflag of the signal "all piston in upper position" to activate hub counter
      Shothub : Bool;   // Piston is metering to make a shot
      Selection_Metering : Bool;   // Request of metering piston, if release is given metring starts
      Selection_Filling : Bool;   // Request of filling piston, if release is given filling starts
      Pos_Weekends_Pause : Bool;   // All pistons are in pause position during manual mode
      Cylinderservice : Bool;   // Key-switch select cylinder service yes/no
      Spare_1_3 : Bool;
      Spare_1_4 : Bool;
      Spare_1_5 : Bool;
      Spare_1_6 : Bool;
      Block_is_active : Bool;   // Function block was passed through // At least 1 piston is active
   END_STRUCT;
END_TYPE

TYPE "UDT062_Cylinder"
TITLE = State of cylinder at piston machine
VERSION : 0.0
   STRUCT
      Metering_runs : Bool;   // Metering piston active
      Filling_runs : Bool;   // Filling piston active
      Release_Metering : Bool;   // Signal release metering of piston present
      Release_Filling : Bool;   // Signal release filling of piston present
      SetValueMetering : Bool;   // Release close loop control metering of piston -> PUC
      SetValueFilling : Bool;   // Release close loop control filling of piston -> PUC
      ReleaseFeedingpump : Bool;   // Release feedpump during filling of piston
      FLT_P_VentingHyd : Bool;   // Fault during depressurizing to vent hydraulic after metering
      FLT_PMax_Component : Bool;   // Fault maximum pressure component exceeded
      FLT_MotorprotectFeedp : Bool;   // Fault supply or motor protection feedpump
      FLT_FeP_Runtime : Bool;   // Fault prepressure piston not reached within 10 sec.
      FLT_L_MinScavenger : Bool;   // Fault level rinsing below min. level
      FLT_FeedpPrepressure : Bool;   // Fault prepressure componente of piston to low
      PistonInUpperPos : Bool;   // Piston at upper endposition
      PistonInButtonPos : Bool;   // Piston at lower endposition
      Puls_QPB : Bool;   // Flag of the signal to switch over to the quick pressure build up
      Valve_Metering : Bool;   // Vavle metering of piston
      Valve_Filling : Bool;   // Vavle filling of piston
      Valve_Suction : Bool;   // Vavle at suction side componente of piston
      Valve_ReleaseFilling : Bool;   // Valve release filling of piston
      Valve_VentingHydr : Bool;   // Valve venting hydraulic
      FLT_MaxPresHydraulic : Bool;   // Fault maximum pressure hydraulic at pistonmotion exceeded
      FLT_Packungsueberwachung : Bool;   // Fault Packungs- pressure exceeded during filling of piston
      Block_is_active : Bool;   // Function block cycling // At least 1 piston is active
      Stepnumber : Byte;   // Stepmemory of control during filling and metering
      FLT_CylinderEmptyShot : Bool;   // Fault Piston empty before foaming end
      FLT_LimitSwitch : Bool;   // Fault limit switch component piston defective (upper- , lower position)
      Spare42 : Bool;
      Spare43 : Bool;
      Spare44 : Bool;
      Spare45 : Bool;
      Spare46 : Bool;
      Spare47 : Bool;
   END_STRUCT;
END_TYPE

TYPE "SZL-IDW#16#xy96_Header"
VERSION : 0.1
   STRUCT
      SZL_ID : Word;
      INDEX : Word;
      LENTHDR : Int;
      N_DR : Int;
   END_STRUCT;
END_TYPE

TYPE "TransmittingError"
VERSION : 0.1
   STRUCT
      Address : Hw_Io;
      Index : Int;
      Length : Int;
      State : DWord;
   END_STRUCT;
END_TYPE

TYPE "UDT014_LP_Circulation_MH"
VERSION : 0.1
   STRUCT
      Flag_Counter : Bool;
      Red_Circulation_On : Bool;
      Start_Flushing : Bool;
      Single_SWU : Bool;
      Change_cycle : Bool;
      Reserve05 : Bool;
      Reserve06 : Bool;
      Reserve07 : Bool;
      Reserve08 : Bool;
      Reserve09 : Bool;
      Reserve10 : Bool;
      Reserve11 : Bool;
      Reserve12 : Bool;
      Reserve13 : Bool;
      Reserve14 : Bool;
      Reserve15 : Bool;
      Amount_MH_for_LP_Circ : Int;
      MH_flushing_finished : Int;
      Reserve16 : Int;
      Reserve17 : Int;
   END_STRUCT;
END_TYPE

